// TIA Portal project "manf386lab6" (V16)

(* hardware
DEVICE "S71500/ET200MP station_1"  S7-1500 station
   slot 0: "Rail_0"  Rack  6ES7 590-1***0-0AA0
   slot 1: "a0"  CPU 1512C-1 PN  6ES7 512-1CK01-0AB0  V2.8
      slot 3: "CPU display_1"  6ES7591-1AA00-0AA0
      slot 32768: "PROFINET interface_1"  X1
         slot 32769: "Port_1"  X1 P1
         slot 32770: "Port_2"  X1 P2
      slot 34817: "Virtual CP interface port_1"  Virtual CP interface port  Virtual CP interface port
DEVICE "MPS distribution touchscreen"  KTP700 Basic PN
   slot 0: "MPS distribution touchscreen"  KTP700 Basic PN  6AV2 123-2GB03-0AX0  16.0.0.0
   slot 1: "HMI_RT_1"  KTP700 Basic PN  6AV2 123-2GB03-0AX0  16.0.0.0
   slot 5: "MPS distribution touchscreen.IE_CP_1"  PROFINET Interface  16.0.0.0
      slot 1: "PROFINET Interface_1"  PROFINET Interface
         slot 1: "Port_1"  Port
*)

// ===== PLC "a0"  CPU 1512C-1 PN =====

VAR_GLOBAL   // PLC tag table "Default tag table"
   "conv_start_I" AT %I10.0 : Bool;   // Workpiece at conveyor start (G1BG1)
   "conv_center_I" AT %I10.1 : Bool;   // Workpiece at conveyor center (G1BG2)
   "conv_end_I" AT %I10.2 : Bool;   // Workpiece NOT at conveyor end (G1BG3)
   "start" AT %I11.0 : Bool;   // Start button
   "stop" AT %I11.1 : Bool;   // Stop Button (NC)
   "key" AT %I11.2 : Bool;   // Key switch (auto/man) (horizontal is true)
   "reset" AT %I11.3 : Bool;   // Reset button
   "panel_I6" AT %I11.6 : Bool;   // Control panel I6
   "panel_I7" AT %I11.7 : Bool;   // Control panel I7
   "conv_fwd" AT %Q4.0 : Bool;   // Conveyor motor forward (G1MA1)
   "conv_bwd" AT %Q4.1 : Bool;   // Conveyor motor backward (G1MA1)
   "retract_gate_Q" AT %Q4.3 : Bool;   // Retract gate (G1MB2)
   "start_LED" AT %Q5.0 : Bool;   // Start indicator light
   "reset_LED" AT %Q5.1 : Bool;   // Reset indicator light
   "Q1_LED" AT %Q5.2 : Bool;   // Indicator light Q1
   "Q2_LED" AT %Q5.3 : Bool;   // Indicator light Q2
   "panel_Q4" AT %Q5.4 : Bool;   // Control panel Q4
   "panel_Q5" AT %Q5.5 : Bool;   // Control panel Q5
   "panel_Q6" AT %Q5.6 : Bool;   // Control panel Q6
   "panel_Q7" AT %Q5.7 : Bool;   // Control panel Q7
   "slide_retracted_I" AT %I10.4 : Bool;   // Slide retracted (C2BG1)
   "slide_extended_I" AT %I10.5 : Bool;   // Slide extended (C2BG2)
   "magazine_empty" AT %I10.6 : Bool;   // Magazine empty (C2BG3)
   "separator" AT %Q4.2 : Bool;   // Extend separator (G1MB1)
   "slide_extend_Q" AT %Q4.4 : Bool;   // Extend slide (C2MB1)
   "main_task_en" AT %Q4.5 : Bool;
   "stop_main_task" AT %Q4.6 : Bool;
END_VAR

DATA_BLOCK "Main [OB1]_DB"   // DB1
{ S7_Optimized_Access := 'TRUE' }
VERSION : 0.1
// stored: InstanceOfName Main [OB1]
"Main [OB1]"
BEGIN
END_DATA_BLOCK

DATA_BLOCK "Block_1_DB"   // DB2
{ S7_Optimized_Access := 'TRUE' }
VERSION : 0.1
// stored: InstanceOfName Block_1
"Block_1"
BEGIN
END_DATA_BLOCK

DATA_BLOCK "HMI Communication"   // DB3
{ S7_Optimized_Access := 'TRUE' }
VERSION : 0.1
   VAR
      conv_start_I : Bool;   // Workpiece at conveyor start (G1BG1)
      conv_center_I : Bool;   // Workpiece at conveyor center (G1BG2)
      conv_end_I : Bool;   // Workpiece NOT at conveyor end (G1BG3)
      start : Bool;   // Start button
      stop : Bool;   // Stop Button (NC)
      key : Bool;   // Key switch (auto/man) (horizontal is true)
      reset : Bool;   // Reset button
      panel_I6 : Bool;   // Control panel I6
      panel_I7 : Bool;   // Control panel I7
      conv_fwd : Bool;   // Conveyor motor forward (G1MA1)
      conv_bwd : Bool;   // Conveyor motor backward (G1MA1)
      retract_gate_Q : Bool;   // Retract gate (G1MB2)
      start_LED : Bool;   // Start indicator light
      reset_LED : Bool;   // Reset indicator light
      Q1_LED : Bool;   // Indicator light Q1
      Q2_LED : Bool;   // Indicator light Q2
      panel_Q4 : Bool;   // Control panel Q4
      panel_Q5 : Bool;   // Control panel Q5
      panel_Q6 : Bool;   // Control panel Q6
      panel_Q7 : Bool;   // Control panel Q7
      slide_retracted_I : Bool;   // Slide retracted (C2BG1)
      slide_extended_I : Bool;   // Slide extended (C2BG2)
      magazine_empty : Bool;   // Magazine empty (C2BG3)
      separator : Bool;   // Extend separator (G1MB1)
      slide_extend_Q : Bool;   // Extend slide (C2MB1)
      main_task_en : Bool;
      stop_main_task : Bool;
   END_VAR
BEGIN
END_DATA_BLOCK

FUNCTION_BLOCK "Main [OB1]"   // FB1, GRAPH_PLUS
{ S7_Optimized_Access := 'TRUE' }
VERSION : 0.1
   VAR_INPUT
      OFF_SQ : Bool := false;   // Turn sequence off
      INIT_SQ : Bool := false;   // Set sequence to initial state
      ACK_EF : Bool := false;   // Acknowledge all errors and faults
      S_PREV : Bool := false;   // Output previous step in parameter S_NO
      S_NEXT : Bool := false;   // Indicate next step in parameter S_NO
      SW_AUTO : Bool := false;   // Automatic mode
      SW_TAP : Bool := false;   // Semiautomatic/switch with transition
      SW_TOP : Bool := false;   // Semiautomatic/ignore transition
      SW_MAN : Bool := false;   // Manual mode
      S_SEL : Int := 0;   // Select step to be output to S_NO
      S_ON : Bool := false;   // Activate step indicated in S_NO
      S_OFF : Bool := false;   // Deactivate step indicated S_NO
      T_PUSH : Bool := false;   // Enable transition to switch in semi automatic mode
   END_VAR
   VAR_OUTPUT
      S_NO : Int := 0;   // Step number
      S_MORE : Bool := false;   // More steps are available and can be shown in S_NO
      S_ACTIVE : Bool := false;   // Step indicated in S_NO is active
      ERR_FLT : Bool := false;   // Interlock or supervision group error
      AUTO_ON : Bool := false;   // Automatic mode is active
      TAP_ON : Bool := false;   // Semiautomatic mode/step with transition enabled
      TOP_ON : Bool := false;   // Semiautomatic mode/ignore transition enabled
      MAN_ON : Bool := false;   // Manual mode is active
   END_VAR
   VAR
      HMI_INFO : Array[0..8] of UInt;
      IF_PAR : G7_IfParPlus_V6;
      RT_DATA : G7_RTDataPlus_V6;   // Internal data area
      key : G7_TransitionPlus_V6;   // Transition structure
      reset_button : G7_TransitionPlus_V6;   // Transition structure
      start_button : G7_TransitionPlus_V6;   // Transition structure
      "stop/man" : G7_TransitionPlus_V6;   // Transition structure
      nan1 : G7_StepPlus_V6;   // Step structure
      reset_led : G7_StepPlus_V6;   // Step structure
      waitForStart : G7_StepPlus_V6;   // Step structure
      "main task" : G7_StepPlus_V6;   // Step structure
      SINI : Array[0..1] of USInt;
      LSTT : Array[0..3] of USInt;
      ATAJ : Array[0..3] of USInt;
      ATAB : Array[0..3] of USInt;
      PSTT : Array[0..3] of USInt;
      NSTT : Array[0..3] of USInt;
      ASSJ : Array[0..3] of USInt;
      ASSB : Array[0..3] of USInt;
      PTTS : Array[0..3] of USInt;
      NTTS : Array[0..3] of USInt;
      SW_SQTS : Array[0..3] of USInt;
      SWITCH : Array[0..0] of USInt;
      TVX : Array[0..1] of USInt;
      TTX : Array[0..1] of USInt;
      TSX : Array[0..1] of USInt;
      S00X : Array[0..1] of USInt;
      SOFFX : Array[0..1] of USInt;
      SONX : Array[0..1] of USInt;
      SAX : Array[0..1] of USInt;
      SERRX : Array[0..4] of USInt;
      SMX : Array[0..4] of USInt;
      S0X : Array[0..4] of USInt;
      S1X : Array[0..4] of USInt;
      IL_ALARM_INST : Diag_Alarm;
      SUP_ALARM_INST : Diag_Alarm;
      STEP_TIME_ALARM_INST : Diag_Alarm;
      IEC_TIMER_INST : IEC_TIMER;
      TRANSACTION_FLAG : Bool := false;
   END_VAR
   VAR_TEMP
      main_task_en : Bool;
   END_VAR
   // SINI[0] := 2;
   // LSTT[0] := 255;
   // LSTT[1] := 255;
   // LSTT[2] := 255;
   // LSTT[3] := 1;
   // ATAJ[1] := 1;
   // ATAJ[2] := 2;
   // ATAJ[3] := 3;
   // ATAB[1] := 1;
   // ATAB[2] := 2;
   // ATAB[3] := 3;
   // PSTT[1] := 1;
   // PSTT[2] := 2;
   // PSTT[3] := 3;
   // NSTT[0] := 1;
   // NSTT[1] := 2;
   // NSTT[2] := 3;
   // NSTT[3] := 1;
   // ASSJ[1] := 1;
   // ASSJ[2] := 2;
   // ASSJ[3] := 3;
   // ASSB[1] := 1;
   // ASSB[2] := 2;
   // ASSB[3] := 3;
   // PTTS[0] := 255;
   // PTTS[2] := 1;
   // PTTS[3] := 2;
   // NTTS[1] := 1;
   // NTTS[2] := 2;
   // NTTS[3] := 3;
   // TVX[0] := 16#1;
   // TTX[0] := 16#1;
   // TSX[0] := 16#1;
   // S00X[0] := 16#1;
   // SOFFX[0] := 16#1;
   // SONX[0] := 16#1;
   // SAX[0] := 16#1;
   // SERRX[0] := 16#1;
   // SMX[0] := 16#1;
   // S0X[0] := 16#1;
   // S1X[0] := 16#1;
BEGIN
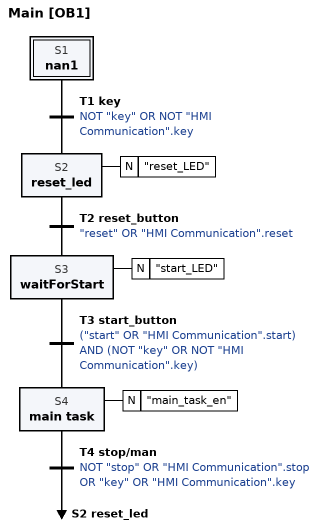
   // sequencer 1
   INITIAL_STEP nan1:   // S1, max time T#10S, warning time T#7S
   END_STEP
   TRANSITION key FROM nan1 TO reset_led   // T1
      := NOT "key" OR NOT "HMI Communication".key;
   END_TRANSITION
   STEP reset_led:   // S2, max time T#10S, warning time T#7S
              N    "reset_LED"
   END_STEP
   TRANSITION reset_button FROM reset_led TO waitForStart   // T2
      := "reset" OR "HMI Communication".reset;
   END_TRANSITION
   STEP waitForStart:   // S3, max time T#10S, warning time T#7S
              N    "start_LED"
   END_STEP
   TRANSITION start_button FROM waitForStart TO "main task"   // T3
      := ("start" OR "HMI Communication".start) AND (NOT "key" OR NOT "HMI Communication".key);
   END_TRANSITION
   STEP "main task":   // S4, max time T#10S, warning time T#7S
              N    "main_task_en"
   END_STEP
   TRANSITION "stop/man" FROM "main task" TO reset_led   // T4, jump
      := NOT "stop" OR "HMI Communication".stop OR "key" OR "HMI Communication".key;
   END_TRANSITION
END_FUNCTION_BLOCK

FUNCTION_BLOCK "Block_1"   // FB2, GRAPH_PLUS
{ S7_Optimized_Access := 'TRUE' }
VERSION : 0.1
   VAR_INPUT
      OFF_SQ : Bool := false;   // Turn sequence off
      INIT_SQ : Bool := false;   // Set sequence to initial state
      ACK_EF : Bool := false;   // Acknowledge all errors and faults
      S_PREV : Bool := false;   // Output previous step in parameter S_NO
      S_NEXT : Bool := false;   // Indicate next step in parameter S_NO
      SW_AUTO : Bool := false;   // Automatic mode
      SW_TAP : Bool := false;   // Semiautomatic/switch with transition
      SW_TOP : Bool := false;   // Semiautomatic/ignore transition
      SW_MAN : Bool := false;   // Manual mode
      S_SEL : Int := 0;   // Select step to be output to S_NO
      S_ON : Bool := false;   // Activate step indicated in S_NO
      S_OFF : Bool := false;   // Deactivate step indicated S_NO
      T_PUSH : Bool := false;   // Enable transition to switch in semi automatic mode
   END_VAR
   VAR_OUTPUT
      S_NO : Int := 0;   // Step number
      S_MORE : Bool := false;   // More steps are available and can be shown in S_NO
      S_ACTIVE : Bool := false;   // Step indicated in S_NO is active
      ERR_FLT : Bool := false;   // Interlock or supervision group error
      AUTO_ON : Bool := false;   // Automatic mode is active
      TAP_ON : Bool := false;   // Semiautomatic mode/step with transition enabled
      TOP_ON : Bool := false;   // Semiautomatic mode/ignore transition enabled
      MAN_ON : Bool := false;   // Manual mode is active
   END_VAR
   VAR
      HMI_INFO : Array[0..8] of UInt;
      IF_PAR : G7_IfParPlus_V6;
      RT_DATA : G7_RTDataPlus_V6;   // Internal data area
      pDetected : G7_TransitionPlus_V6;   // Transition structure
      pPrime : G7_TransitionPlus_V6;   // Transition structure
      pFin : G7_TransitionPlus_V6;   // Transition structure
      pWait : G7_StepPlus_V6;   // Step structure
      pPushMid : G7_StepPlus_V6;   // Step structure
      sPushEnd : G7_StepPlus_V6;   // Step structure
      SINI : Array[0..1] of USInt;
      LSTT : Array[0..2] of USInt;
      ATAJ : Array[0..2] of USInt;
      ATAB : Array[0..2] of USInt;
      PSTT : Array[0..2] of USInt;
      NSTT : Array[0..2] of USInt;
      ASSJ : Array[0..2] of USInt;
      ASSB : Array[0..2] of USInt;
      PTTS : Array[0..2] of USInt;
      NTTS : Array[0..2] of USInt;
      SW_SQTS : Array[0..2] of USInt;
      SWITCH : Array[0..0] of USInt;
      TVX : Array[0..1] of USInt;
      TTX : Array[0..1] of USInt;
      TSX : Array[0..1] of USInt;
      S00X : Array[0..1] of USInt;
      SOFFX : Array[0..1] of USInt;
      SONX : Array[0..1] of USInt;
      SAX : Array[0..1] of USInt;
      SERRX : Array[0..3] of USInt;
      SMX : Array[0..3] of USInt;
      S0X : Array[0..3] of USInt;
      S1X : Array[0..3] of USInt;
      IL_ALARM_INST : Diag_Alarm;
      SUP_ALARM_INST : Diag_Alarm;
      STEP_TIME_ALARM_INST : Diag_Alarm;
      IEC_TIMER_INST : IEC_TIMER;
      TRANSACTION_FLAG : Bool := false;
   END_VAR
   // SINI[0] := 2;
   // LSTT[0] := 255;
   // LSTT[1] := 255;
   // ATAJ[1] := 1;
   // ATAJ[2] := 2;
   // ATAB[1] := 1;
   // ATAB[2] := 2;
   // PSTT[1] := 1;
   // PSTT[2] := 2;
   // NSTT[0] := 1;
   // NSTT[1] := 2;
   // ASSJ[1] := 1;
   // ASSJ[2] := 2;
   // ASSB[1] := 1;
   // ASSB[2] := 2;
   // PTTS[0] := 255;
   // PTTS[2] := 1;
   // NTTS[1] := 1;
   // NTTS[2] := 2;
   // TVX[0] := 16#1;
   // TTX[0] := 16#1;
   // TSX[0] := 16#1;
   // S00X[0] := 16#1;
   // SOFFX[0] := 16#1;
   // SONX[0] := 16#1;
   // SAX[0] := 16#1;
   // SERRX[0] := 16#1;
   // SMX[0] := 16#1;
   // S0X[0] := 16#1;
   // S1X[0] := 16#1;
BEGIN
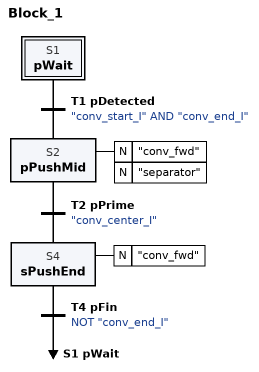
   // sequencer 1
   INITIAL_STEP pWait:   // S1, max time T#10S, warning time T#7S
   END_STEP
   TRANSITION pDetected FROM pWait TO pPushMid   // T1
      := "conv_start_I" AND "conv_end_I";
   END_TRANSITION
   STEP pPushMid:   // S2, max time T#10S, warning time T#7S
              N    "conv_fwd"
              N    "separator"
   END_STEP
   TRANSITION pPrime FROM pPushMid TO sPushEnd   // T2
      := "conv_center_I";
   END_TRANSITION
   STEP sPushEnd:   // S4, max time T#10S, warning time T#7S
              N    "conv_fwd"
   END_STEP
   TRANSITION pFin FROM sPushEnd TO pWait   // T4, jump
      := NOT "conv_end_I";
   END_TRANSITION
END_FUNCTION_BLOCK

ORGANIZATION_BLOCK "Main LAD"   // OB1, LAD, ProgramCycle
TITLE = "Main Program Sweep (Cycle)"
{ S7_Optimized_Access := 'TRUE' }
VERSION : 0.1
   VAR_INPUT
      Initial_Call : Bool;   // Initial call of this OB
      Remanence : Bool;   // =True, if remanent data are available
   END_VAR
   VAR_TEMP
      main_task_running : Bool;
      Temp_2 : Bool;
   END_VAR
BEGIN

REGION Network 1
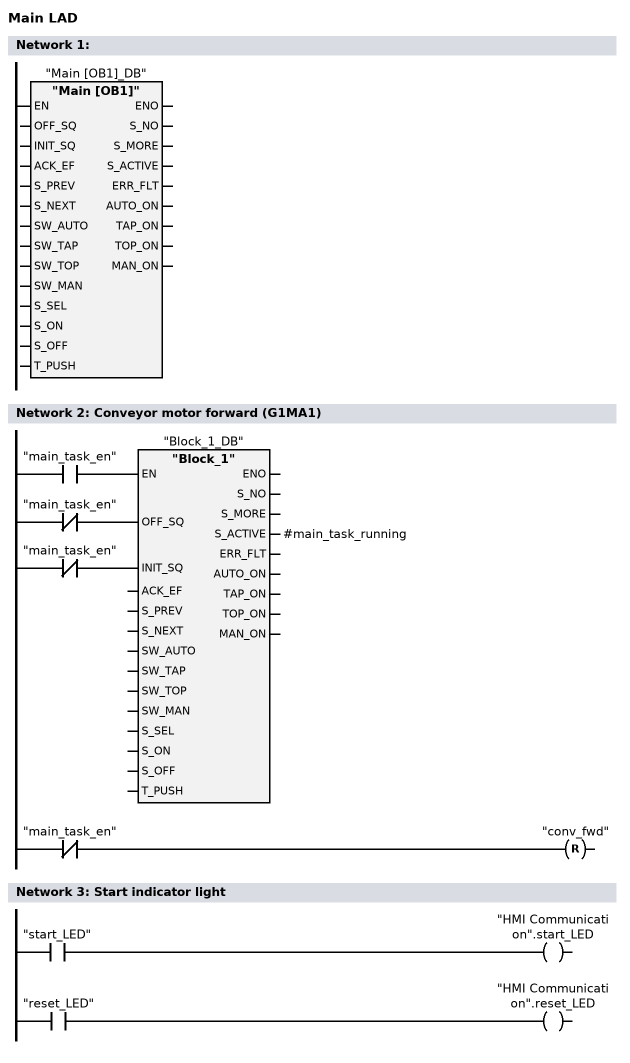
   RUNG wire#powerrail
      "Main [OB1]_DB"(OFF_SQ :=, INIT_SQ :=, ACK_EF :=, S_PREV :=, S_NEXT :=, SW_AUTO :=, SW_TAP :=, SW_TOP :=, SW_MAN :=, S_SEL :=, S_ON :=, S_OFF :=, T_PUSH :=, S_NO =>, S_MORE =>, S_ACTIVE =>, ERR_FLT =>, AUTO_ON =>, TAP_ON =>, TOP_ON =>, MAN_ON =>)
   END_RUNG
   // the same network as SCL:
   "Main [OB1]_DB"();   // "Main [OB1]"
END_REGION

REGION Network 2: Conveyor motor forward (G1MA1)
   RUNG wire#powerrail
      Contact( "main_task_en" )
      "Block_1_DB"(OFF_SQ := wire#w1, INIT_SQ := wire#w2, ACK_EF :=, S_PREV :=, S_NEXT :=, SW_AUTO :=, SW_TAP :=, SW_TOP :=, SW_MAN :=, S_SEL :=, S_ON :=, S_OFF :=, T_PUSH :=, S_NO =>, S_MORE =>, S_ACTIVE => #main_task_running, ERR_FLT =>, AUTO_ON =>, TAP_ON =>, TOP_ON =>, MAN_ON =>)
   END_RUNG
   RUNG wire#powerrail
      I_Contact( "main_task_en" )
   END_RUNG wire#w1
   RUNG wire#powerrail
      I_Contact( "main_task_en" )
   END_RUNG wire#w2
   RUNG wire#powerrail
      I_Contact( "main_task_en" )
      R_Coil( "conv_fwd" )
   END_RUNG
   // the same network as SCL:
   IF "main_task_en" THEN
       "Block_1_DB"(OFF_SQ := NOT "main_task_en", INIT_SQ := NOT "main_task_en", S_ACTIVE => #main_task_running);   // "Block_1"
   END_IF;
   IF NOT "main_task_en" THEN "conv_fwd" := FALSE; END_IF;
END_REGION

REGION Network 3: Start indicator light
   RUNG wire#powerrail
      Contact( "start_LED" )
      Coil( "HMI Communication".start_LED )
   END_RUNG
   RUNG wire#powerrail
      Contact( "reset_LED" )
      Coil( "HMI Communication".reset_LED )
   END_RUNG
   // the same network as SCL:
   "HMI Communication".start_LED := "start_LED";
   "HMI Communication".reset_LED := "reset_LED";
END_REGION
END_ORGANIZATION_BLOCK

(* ===== HMI "HMI_RT_1" =====
system functions are stored by id; their names below are inferred from use
connection "HMI_Connection_1": ETHERNET, SMART_S7_1500_OMS

HMI tags "Default tag table"
   "HMI Communication_start" : Bool = PLC "HMI Communication".start, 100 ms
   "HMI Communication_stop" : Bool = PLC "HMI Communication".stop, 100 ms
   "HMI Communication_reset" : Bool = PLC "HMI Communication".reset, 100 ms
   "HMI Communication_start_LED" : Bool = PLC "HMI Communication".start_LED, 100 ms
   "HMI Communication_reset_LED" : Bool = PLC "HMI Communication".reset_LED, 100 ms
   "HMI Communication_key" : Bool = PLC "HMI Communication".key, 100 ms
   "reset_LED" : Bool = PLC reset_LED AT %Q5.1, 1 s

screen "Screen_1" 800x480
   Button "Button_1" at 48,33 size 236x119; TextOff 'Start'
      on Press: function_b14e0dd5("HMI Communication_start", 0)
   Button "Button_2" at 284,32 size 245x120; TextOff 'Stop'
      on Press: function_b14e0dd5("HMI Communication_stop", 0)
   Button "Button_3" at 529,32 size 240x120; TextOff 'Reset'
      on Press: function_b14e0dd5("HMI Communication_reset", 0)
   Circle "Circle_1" at 56,42 size 48x48
      Appearance <- "HMI Communication_start_LED"
   Circle "Circle_2" at 542,42 size 48x48
      Appearance <- "reset_LED"
   Switch "Switch_1" at 48,316 size 282x95; CaptionText 'Switch'; TextOff 'Auto'; TextOn 'Man'
      ProcessValue <- "HMI Communication_key"
      on SwitchOn: SetBit("HMI Communication_key")
      on SwitchOff: ResetBit("HMI Communication_key")
*)